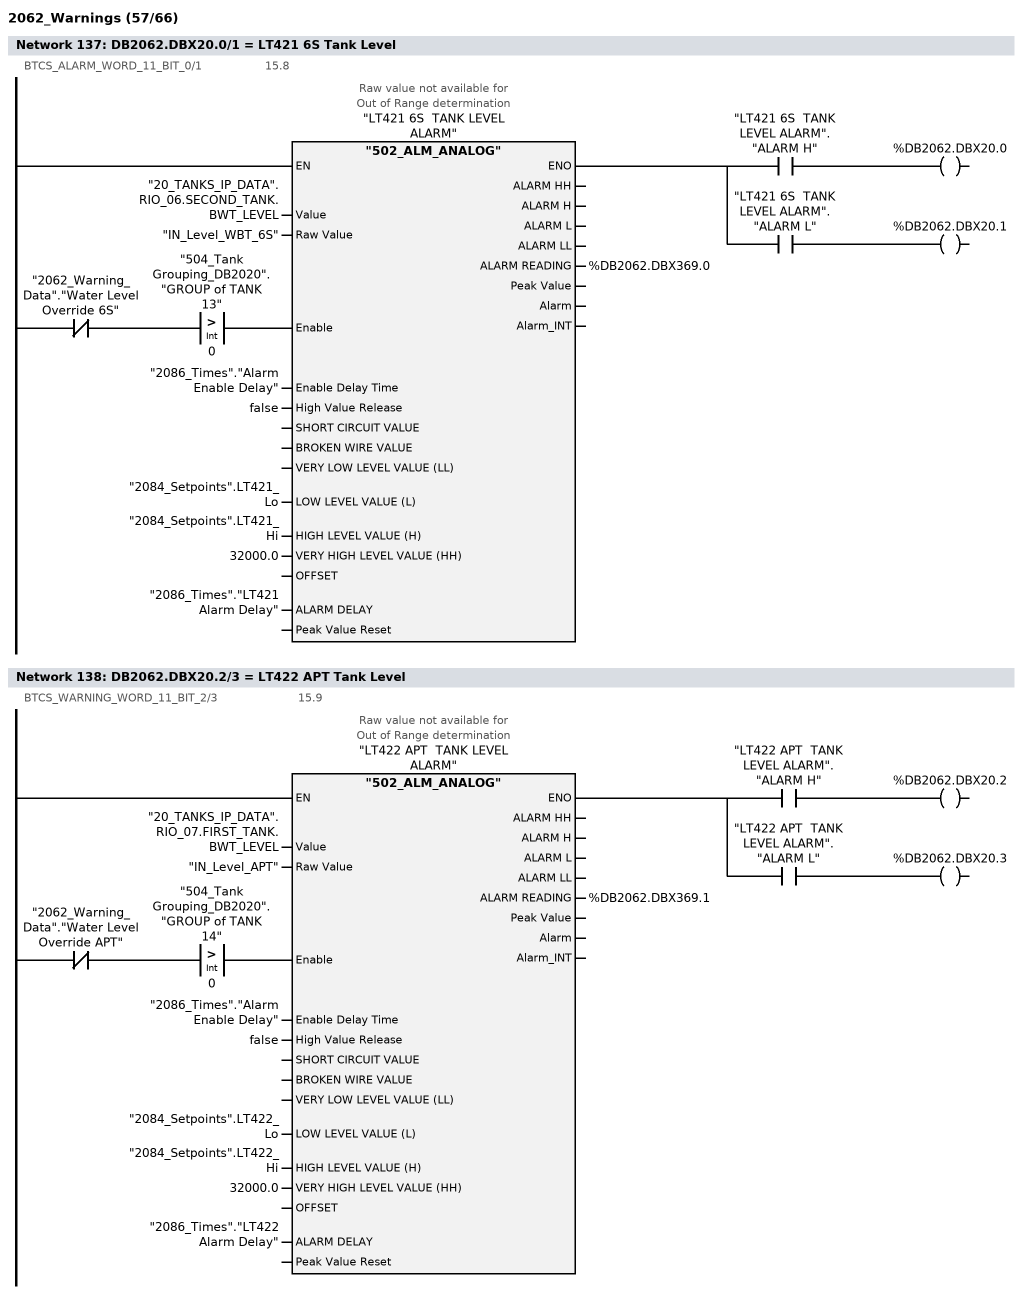
   RUNG wire#powerrail
      "LT421 6S  TANK LEVEL ALARM"(Enable := wire#w1, Value := "20_TANKS_IP_DATA".RIO_06.SECOND_TANK.BWT_LEVEL, "Raw Value" := "IN_Level_WBT_6S", "Enable Delay Time" := "2086_Times"."Alarm Enable Delay", "High Value Release" := false, "SHORT CIRCUIT VALUE" :=, "BROKEN WIRE VALUE" :=, "VERY LOW LEVEL VALUE (LL)" :=, "LOW LEVEL VALUE (L)" := "2084_Setpoints".LT421_Lo, "HIGH LEVEL VALUE (H)" := "2084_Setpoints".LT421_Hi, "VERY HIGH LEVEL VALUE (HH)" := 32000.0, OFFSET :=, "ALARM DELAY" := "2086_Times"."LT421 Alarm Delay", "Peak Value Reset" :=, "ALARM HH" =>, "ALARM H" =>, "ALARM L" =>, "ALARM LL" =>, "ALARM READING" => %DB2062.DBX369.0, "Peak Value" =>, Alarm =>, Alarm_INT =>)   // Raw value not available for Out of Range determination
      wire#w2
      Contact( "LT421 6S  TANK LEVEL ALARM"."ALARM H" )
      Coil( %DB2062.DBX20.0 )
   END_RUNG
   RUNG wire#powerrail
      I_Contact( "2062_Warning_Data"."Water Level Override 6S" )
      { S7_Templates := "SrcType := Int" } GT_Contact(in1 := "504_Tank Grouping_DB2020"."GROUP of TANK 13", in2 := 0)
   END_RUNG wire#w1
   RUNG wire#w2
      Contact( "LT421 6S  TANK LEVEL ALARM"."ALARM L" )
      Coil( %DB2062.DBX20.1 )
   END_RUNG
   // the same network as SCL:
   "LT421 6S  TANK LEVEL ALARM"(Value := "20_TANKS_IP_DATA".RIO_06.SECOND_TANK.BWT_LEVEL,   // "502_ALM_ANALOG": Raw value not available for Out of Range determination
                           "Raw Value" := "IN_Level_WBT_6S",
                           Enable := NOT "2062_Warning_Data"."Water Level Override 6S" AND ("504_Tank Grouping_DB2020"."GROUP of TANK 13" > 0),
                           "Enable Delay Time" := "2086_Times"."Alarm Enable Delay",
                           "High Value Release" := false,
                           "LOW LEVEL VALUE (L)" := "2084_Setpoints".LT421_Lo,
                           "HIGH LEVEL VALUE (H)" := "2084_Setpoints".LT421_Hi,
                           "VERY HIGH LEVEL VALUE (HH)" := 32000.0,
                           "ALARM DELAY" := "2086_Times"."LT421 Alarm Delay",
                           "ALARM READING" => %DB2062.DBX369.0,
                           ENO => #_w1);
   %DB2062.DBX20.0 := #_w1 AND "LT421 6S  TANK LEVEL ALARM"."ALARM H";
   %DB2062.DBX20.1 := #_w1 AND "LT421 6S  TANK LEVEL ALARM"."ALARM L";
END_REGION

REGION Network 138: DB2062.DBX20.2/3 = LT422 APT Tank Level
   // BTCS_WARNING_WORD_11_BIT_2/3                       15.9
   RUNG wire#powerrail
      "LT422 APT  TANK LEVEL ALARM"(Enable := wire#w1, Value := "20_TANKS_IP_DATA".RIO_07.FIRST_TANK.BWT_LEVEL, "Raw Value" := "IN_Level_APT", "Enable Delay Time" := "2086_Times"."Alarm Enable Delay", "High Value Release" := false, "SHORT CIRCUIT VALUE" :=, "BROKEN WIRE VALUE" :=, "VERY LOW LEVEL VALUE (LL)" :=, "LOW LEVEL VALUE (L)" := "2084_Setpoints".LT422_Lo, "HIGH LEVEL VALUE (H)" := "2084_Setpoints".LT422_Hi, "VERY HIGH LEVEL VALUE (HH)" := 32000.0, OFFSET :=, "ALARM DELAY" := "2086_Times"."LT422 Alarm Delay", "Peak Value Reset" :=, "ALARM HH" =>, "ALARM H" =>, "ALARM L" =>, "ALARM LL" =>, "ALARM READING" => %DB2062.DBX369.1, "Peak Value" =>, Alarm =>, Alarm_INT =>)   // Raw value not available for Out of Range determination
      wire#w2
      Contact( "LT422 APT  TANK LEVEL ALARM"."ALARM H" )
      Coil( %DB2062.DBX20.2 )
   END_RUNG
   RUNG wire#powerrail
      I_Contact( "2062_Warning_Data"."Water Level Override APT" )
      { S7_Templates := "SrcType := Int" } GT_Contact(in1 := "504_Tank Grouping_DB2020"."GROUP of TANK 14", in2 := 0)
   END_RUNG wire#w1
   RUNG wire#w2
      Contact( "LT422 APT  TANK LEVEL ALARM"."ALARM L" )
      Coil( %DB2062.DBX20.3 )
   END_RUNG
   // the same network as SCL:
   "LT422 APT  TANK LEVEL ALARM"(Value := "20_TANKS_IP_DATA".RIO_07.FIRST_TANK.BWT_LEVEL,   // "502_ALM_ANALOG": Raw value not available for Out of Range determination
                           "Raw Value" := "IN_Level_APT",
                           Enable := NOT "2062_Warning_Data"."Water Level Override APT" AND ("504_Tank Grouping_DB2020"."GROUP of TANK 14" > 0),
                           "Enable Delay Time" := "2086_Times"."Alarm Enable Delay",
                           "High Value Release" := false,
                           "LOW LEVEL VALUE (L)" := "2084_Setpoints".LT422_Lo,
                           "HIGH LEVEL VALUE (H)" := "2084_Setpoints".LT422_Hi,
                           "VERY HIGH LEVEL VALUE (HH)" := 32000.0,
                           "ALARM DELAY" := "2086_Times"."LT422 Alarm Delay",
                           "ALARM READING" => %DB2062.DBX369.1,
                           ENO => #_w1);
   %DB2062.DBX20.2 := #_w1 AND "LT422 APT  TANK LEVEL ALARM"."ALARM H";
   %DB2062.DBX20.3 := #_w1 AND "LT422 APT  TANK LEVEL ALARM"."ALARM L";
END_REGION

REGION Network 140: Alarm Tank 1
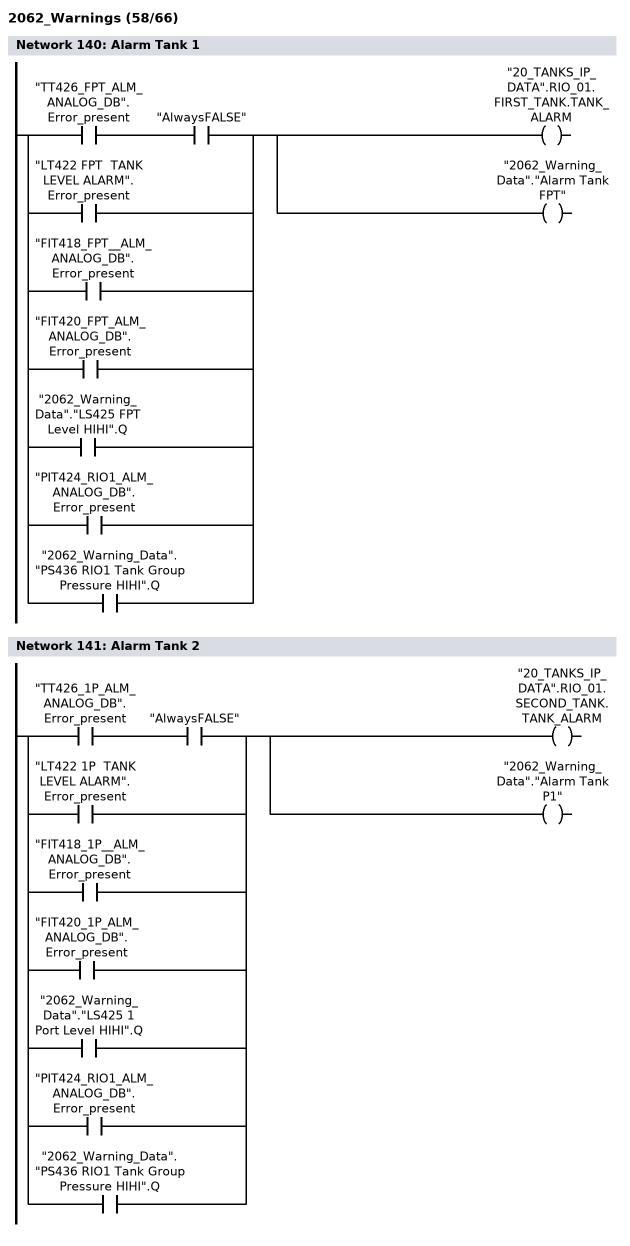
   RUNG wire#powerrail
      Contact( "TT426_FPT_ALM_ANALOG_DB".Error_present )
      Contact( "AlwaysFALSE" )
      wire#w1
      Coil( "20_TANKS_IP_DATA".RIO_01.FIRST_TANK.TANK_ALARM )
   END_RUNG
   RUNG wire#powerrail
      Contact( "LT422 FPT  TANK LEVEL ALARM".Error_present )
   END_RUNG wire#w1
   RUNG wire#powerrail
      Contact( "FIT418_FPT__ALM_ANALOG_DB".Error_present )
   END_RUNG wire#w1
   RUNG wire#powerrail
      Contact( "FIT420_FPT_ALM_ANALOG_DB".Error_present )
   END_RUNG wire#w1
   RUNG wire#powerrail
      Contact( "2062_Warning_Data"."LS425 FPT Level HIHI".Q )
   END_RUNG wire#w1
   RUNG wire#powerrail
      Contact( "PIT424_RIO1_ALM_ANALOG_DB".Error_present )
   END_RUNG wire#w1
   RUNG wire#powerrail
      Contact( "2062_Warning_Data"."PS436 RIO1 Tank Group Pressure HIHI".Q )
   END_RUNG wire#w1
   RUNG wire#w1
      Coil( "2062_Warning_Data"."Alarm Tank FPT" )
   END_RUNG
   // the same network as SCL:
   "20_TANKS_IP_DATA".RIO_01.FIRST_TANK.TANK_ALARM := ("TT426_FPT_ALM_ANALOG_DB".Error_present AND "AlwaysFALSE") OR "LT422 FPT  TANK LEVEL ALARM".Error_present OR "FIT418_FPT__ALM_ANALOG_DB".Error_present OR "FIT420_FPT_ALM_ANALOG_DB".Error_present OR "2062_Warning_Data"."LS425 FPT Level HIHI".Q OR "PIT424_RIO1_ALM_ANALOG_DB".Error_present OR "2062_Warning_Data"."PS436 RIO1 Tank Group Pressure HIHI".Q;
   "2062_Warning_Data"."Alarm Tank FPT" := "20_TANKS_IP_DATA".RIO_01.FIRST_TANK.TANK_ALARM;
END_REGION

REGION Network 141: Alarm Tank 2
   RUNG wire#powerrail
      Contact( "TT426_1P_ALM_ANALOG_DB".Error_present )
      Contact( "AlwaysFALSE" )
      wire#w1
      Coil( "20_TANKS_IP_DATA".RIO_01.SECOND_TANK.TANK_ALARM )
   END_RUNG
   RUNG wire#powerrail
      Contact( "LT422 1P  TANK LEVEL ALARM".Error_present )
   END_RUNG wire#w1
   RUNG wire#powerrail
      Contact( "FIT418_1P__ALM_ANALOG_DB".Error_present )
   END_RUNG wire#w1
   RUNG wire#powerrail
      Contact( "FIT420_1P_ALM_ANALOG_DB".Error_present )
   END_RUNG wire#w1
   RUNG wire#powerrail
      Contact( "2062_Warning_Data"."LS425 1 Port Level HIHI".Q )
   END_RUNG wire#w1
   RUNG wire#powerrail
      Contact( "PIT424_RIO1_ALM_ANALOG_DB".Error_present )
   END_RUNG wire#w1
   RUNG wire#powerrail
      Contact( "2062_Warning_Data"."PS436 RIO1 Tank Group Pressure HIHI".Q )
   END_RUNG wire#w1
   RUNG wire#w1
      Coil( "2062_Warning_Data"."Alarm Tank P1" )
   END_RUNG
   // the same network as SCL:
   "20_TANKS_IP_DATA".RIO_01.SECOND_TANK.TANK_ALARM := ("TT426_1P_ALM_ANALOG_DB".Error_present AND "AlwaysFALSE") OR "LT422 1P  TANK LEVEL ALARM".Error_present OR "FIT418_1P__ALM_ANALOG_DB".Error_present OR "FIT420_1P_ALM_ANALOG_DB".Error_present OR "2062_Warning_Data"."LS425 1 Port Level HIHI".Q OR "PIT424_RIO1_ALM_ANALOG_DB".Error_present OR "2062_Warning_Data"."PS436 RIO1 Tank Group Pressure HIHI".Q;
   "2062_Warning_Data"."Alarm Tank P1" := "20_TANKS_IP_DATA".RIO_01.SECOND_TANK.TANK_ALARM;
END_REGION

REGION Network 142: Alarm Tank 3
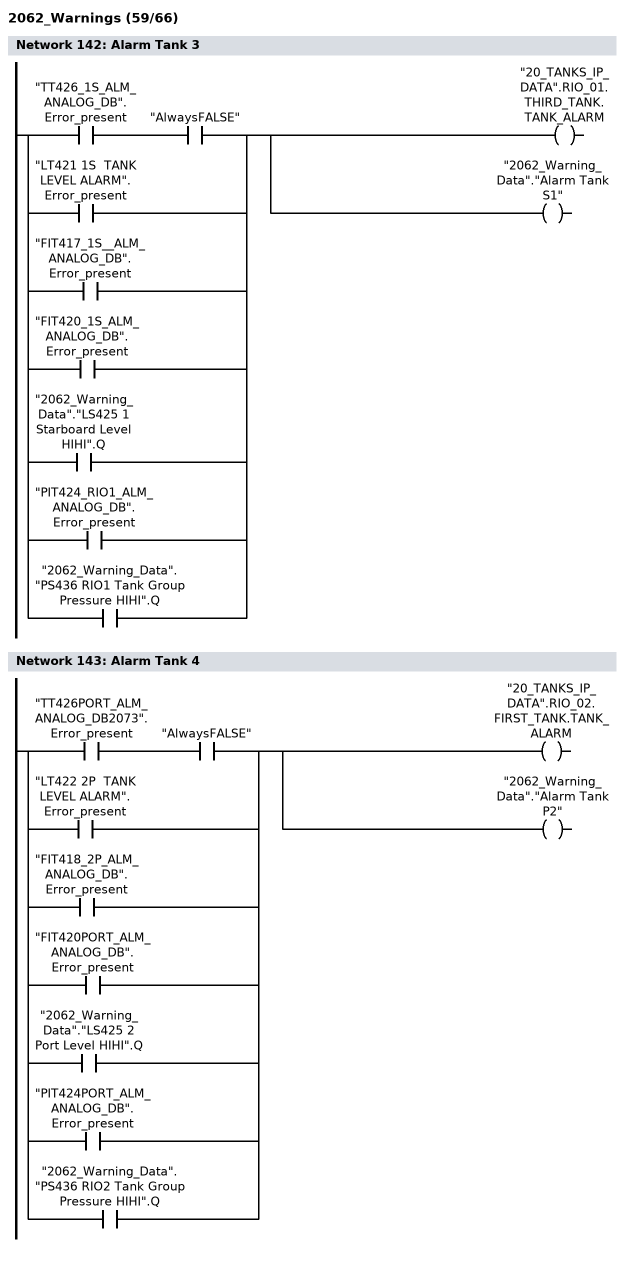
   RUNG wire#powerrail
      Contact( "TT426_1S_ALM_ANALOG_DB".Error_present )
      Contact( "AlwaysFALSE" )
      wire#w1
      Coil( "20_TANKS_IP_DATA".RIO_01.THIRD_TANK.TANK_ALARM )
   END_RUNG
   RUNG wire#powerrail
      Contact( "LT421 1S  TANK LEVEL ALARM".Error_present )
   END_RUNG wire#w1
   RUNG wire#powerrail
      Contact( "FIT417_1S__ALM_ANALOG_DB".Error_present )
   END_RUNG wire#w1
   RUNG wire#powerrail
      Contact( "FIT420_1S_ALM_ANALOG_DB".Error_present )
   END_RUNG wire#w1
   RUNG wire#powerrail
      Contact( "2062_Warning_Data"."LS425 1 Starboard Level HIHI".Q )
   END_RUNG wire#w1
   RUNG wire#powerrail
      Contact( "PIT424_RIO1_ALM_ANALOG_DB".Error_present )
   END_RUNG wire#w1
   RUNG wire#powerrail
      Contact( "2062_Warning_Data"."PS436 RIO1 Tank Group Pressure HIHI".Q )
   END_RUNG wire#w1
   RUNG wire#w1
      Coil( "2062_Warning_Data"."Alarm Tank S1" )
   END_RUNG
   // the same network as SCL:
   "20_TANKS_IP_DATA".RIO_01.THIRD_TANK.TANK_ALARM := ("TT426_1S_ALM_ANALOG_DB".Error_present AND "AlwaysFALSE") OR "LT421 1S  TANK LEVEL ALARM".Error_present OR "FIT417_1S__ALM_ANALOG_DB".Error_present OR "FIT420_1S_ALM_ANALOG_DB".Error_present OR "2062_Warning_Data"."LS425 1 Starboard Level HIHI".Q OR "PIT424_RIO1_ALM_ANALOG_DB".Error_present OR "2062_Warning_Data"."PS436 RIO1 Tank Group Pressure HIHI".Q;
   "2062_Warning_Data"."Alarm Tank S1" := "20_TANKS_IP_DATA".RIO_01.THIRD_TANK.TANK_ALARM;
END_REGION

REGION Network 143: Alarm Tank 4
   RUNG wire#powerrail
      Contact( "TT426PORT_ALM_ANALOG_DB2073".Error_present )
      Contact( "AlwaysFALSE" )
      wire#w1
      Coil( "20_TANKS_IP_DATA".RIO_02.FIRST_TANK.TANK_ALARM )
   END_RUNG
   RUNG wire#powerrail
      Contact( "LT422 2P  TANK LEVEL ALARM".Error_present )
   END_RUNG wire#w1
   RUNG wire#powerrail
      Contact( "FIT418_2P_ALM_ANALOG_DB".Error_present )
   END_RUNG wire#w1
   RUNG wire#powerrail
      Contact( "FIT420PORT_ALM_ANALOG_DB".Error_present )
   END_RUNG wire#w1
   RUNG wire#powerrail
      Contact( "2062_Warning_Data"."LS425 2 Port Level HIHI".Q )
   END_RUNG wire#w1
   RUNG wire#powerrail
      Contact( "PIT424PORT_ALM_ANALOG_DB".Error_present )
   END_RUNG wire#w1
   RUNG wire#powerrail
      Contact( "2062_Warning_Data"."PS436 RIO2 Tank Group Pressure HIHI".Q )
   END_RUNG wire#w1
   RUNG wire#w1
      Coil( "2062_Warning_Data"."Alarm Tank P2" )
   END_RUNG
   // the same network as SCL:
   "20_TANKS_IP_DATA".RIO_02.FIRST_TANK.TANK_ALARM := ("TT426PORT_ALM_ANALOG_DB2073".Error_present AND "AlwaysFALSE") OR "LT422 2P  TANK LEVEL ALARM".Error_present OR "FIT418_2P_ALM_ANALOG_DB".Error_present OR "FIT420PORT_ALM_ANALOG_DB".Error_present OR "2062_Warning_Data"."LS425 2 Port Level HIHI".Q OR "PIT424PORT_ALM_ANALOG_DB".Error_present OR "2062_Warning_Data"."PS436 RIO2 Tank Group Pressure HIHI".Q;
   "2062_Warning_Data"."Alarm Tank P2" := "20_TANKS_IP_DATA".RIO_02.FIRST_TANK.TANK_ALARM;
END_REGION

REGION Network 144: Alarm Tank 5
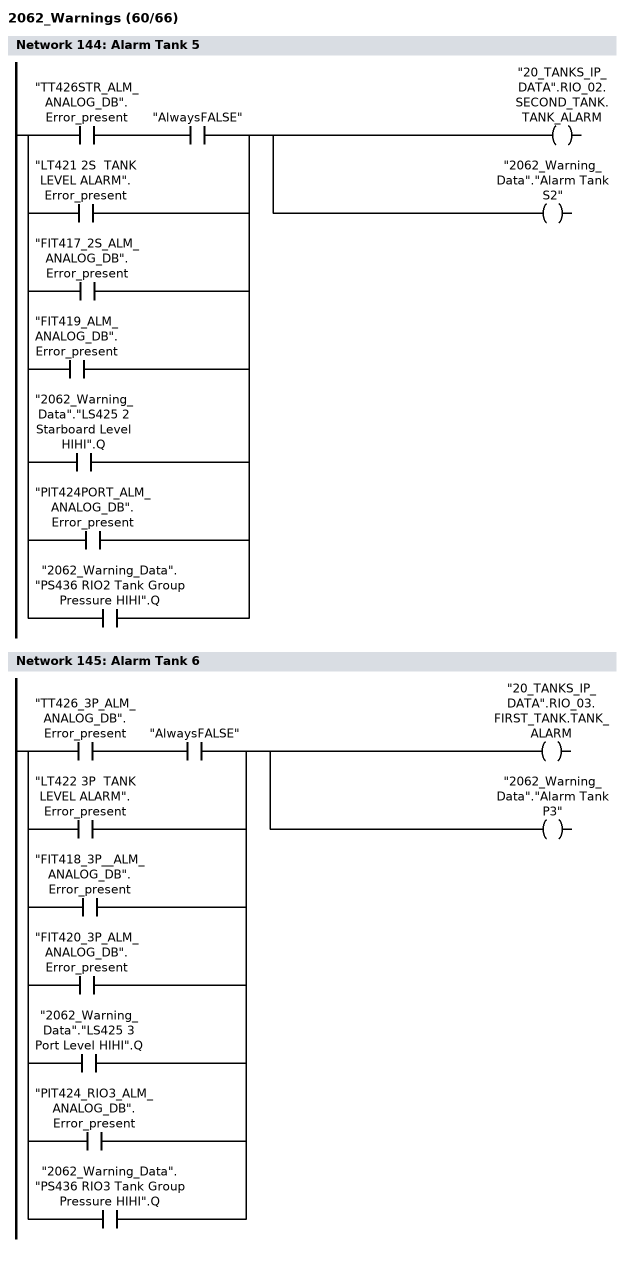
   RUNG wire#powerrail
      Contact( "TT426STR_ALM_ANALOG_DB".Error_present )
      Contact( "AlwaysFALSE" )
      wire#w1
      Coil( "20_TANKS_IP_DATA".RIO_02.SECOND_TANK.TANK_ALARM )
   END_RUNG
   RUNG wire#powerrail
      Contact( "LT421 2S  TANK LEVEL ALARM".Error_present )
   END_RUNG wire#w1
   RUNG wire#powerrail
      Contact( "FIT417_2S_ALM_ANALOG_DB".Error_present )
   END_RUNG wire#w1
   RUNG wire#powerrail
      Contact( "FIT419_ALM_ANALOG_DB".Error_present )
   END_RUNG wire#w1
   RUNG wire#powerrail
      Contact( "2062_Warning_Data"."LS425 2 Starboard Level HIHI".Q )
   END_RUNG wire#w1
   RUNG wire#powerrail
      Contact( "PIT424PORT_ALM_ANALOG_DB".Error_present )
   END_RUNG wire#w1
   RUNG wire#powerrail
      Contact( "2062_Warning_Data"."PS436 RIO2 Tank Group Pressure HIHI".Q )
   END_RUNG wire#w1
   RUNG wire#w1
      Coil( "2062_Warning_Data"."Alarm Tank S2" )
   END_RUNG
   // the same network as SCL:
   "20_TANKS_IP_DATA".RIO_02.SECOND_TANK.TANK_ALARM := ("TT426STR_ALM_ANALOG_DB".Error_present AND "AlwaysFALSE") OR "LT421 2S  TANK LEVEL ALARM".Error_present OR "FIT417_2S_ALM_ANALOG_DB".Error_present OR "FIT419_ALM_ANALOG_DB".Error_present OR "2062_Warning_Data"."LS425 2 Starboard Level HIHI".Q OR "PIT424PORT_ALM_ANALOG_DB".Error_present OR "2062_Warning_Data"."PS436 RIO2 Tank Group Pressure HIHI".Q;
   "2062_Warning_Data"."Alarm Tank S2" := "20_TANKS_IP_DATA".RIO_02.SECOND_TANK.TANK_ALARM;
END_REGION

REGION Network 145: Alarm Tank 6
   RUNG wire#powerrail
      Contact( "TT426_3P_ALM_ANALOG_DB".Error_present )
      Contact( "AlwaysFALSE" )
      wire#w1
      Coil( "20_TANKS_IP_DATA".RIO_03.FIRST_TANK.TANK_ALARM )
   END_RUNG
   RUNG wire#powerrail
      Contact( "LT422 3P  TANK LEVEL ALARM".Error_present )
   END_RUNG wire#w1
   RUNG wire#powerrail
      Contact( "FIT418_3P__ALM_ANALOG_DB".Error_present )
   END_RUNG wire#w1
   RUNG wire#powerrail
      Contact( "FIT420_3P_ALM_ANALOG_DB".Error_present )
   END_RUNG wire#w1
   RUNG wire#powerrail
      Contact( "2062_Warning_Data"."LS425 3 Port Level HIHI".Q )
   END_RUNG wire#w1
   RUNG wire#powerrail
      Contact( "PIT424_RIO3_ALM_ANALOG_DB".Error_present )
   END_RUNG wire#w1
   RUNG wire#powerrail
      Contact( "2062_Warning_Data"."PS436 RIO3 Tank Group Pressure HIHI".Q )
   END_RUNG wire#w1
   RUNG wire#w1
      Coil( "2062_Warning_Data"."Alarm Tank P3" )
   END_RUNG
   // the same network as SCL:
   "20_TANKS_IP_DATA".RIO_03.FIRST_TANK.TANK_ALARM := ("TT426_3P_ALM_ANALOG_DB".Error_present AND "AlwaysFALSE") OR "LT422 3P  TANK LEVEL ALARM".Error_present OR "FIT418_3P__ALM_ANALOG_DB".Error_present OR "FIT420_3P_ALM_ANALOG_DB".Error_present OR "2062_Warning_Data"."LS425 3 Port Level HIHI".Q OR "PIT424_RIO3_ALM_ANALOG_DB".Error_present OR "2062_Warning_Data"."PS436 RIO3 Tank Group Pressure HIHI".Q;
   "2062_Warning_Data"."Alarm Tank P3" := "20_TANKS_IP_DATA".RIO_03.FIRST_TANK.TANK_ALARM;
END_REGION

REGION Network 146: Alarm Tank 7
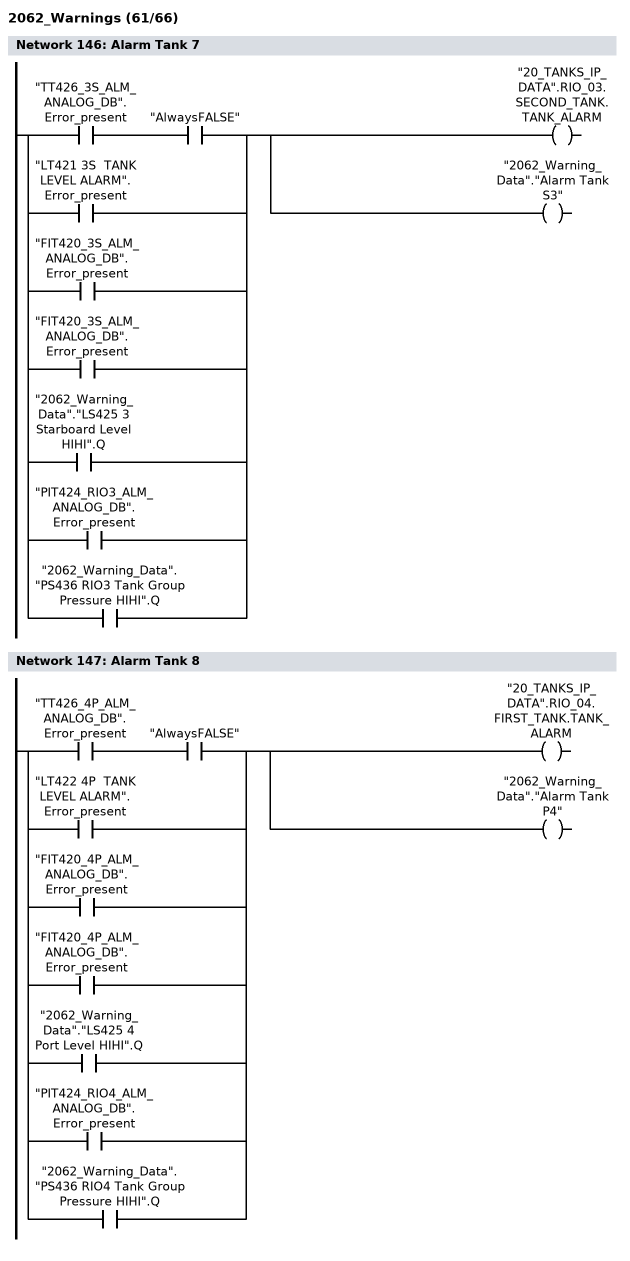
   RUNG wire#powerrail
      Contact( "TT426_3S_ALM_ANALOG_DB".Error_present )
      Contact( "AlwaysFALSE" )
      wire#w1
      Coil( "20_TANKS_IP_DATA".RIO_03.SECOND_TANK.TANK_ALARM )
   END_RUNG
   RUNG wire#powerrail
      Contact( "LT421 3S  TANK LEVEL ALARM".Error_present )
   END_RUNG wire#w1
   RUNG wire#powerrail
      Contact( "FIT420_3S_ALM_ANALOG_DB".Error_present )
   END_RUNG wire#w1
   RUNG wire#powerrail
      Contact( "FIT420_3S_ALM_ANALOG_DB".Error_present )
   END_RUNG wire#w1
   RUNG wire#powerrail
      Contact( "2062_Warning_Data"."LS425 3 Starboard Level HIHI".Q )
   END_RUNG wire#w1
   RUNG wire#powerrail
      Contact( "PIT424_RIO3_ALM_ANALOG_DB".Error_present )
   END_RUNG wire#w1
   RUNG wire#powerrail
      Contact( "2062_Warning_Data"."PS436 RIO3 Tank Group Pressure HIHI".Q )
   END_RUNG wire#w1
   RUNG wire#w1
      Coil( "2062_Warning_Data"."Alarm Tank S3" )
   END_RUNG
   // the same network as SCL:
   "20_TANKS_IP_DATA".RIO_03.SECOND_TANK.TANK_ALARM := ("TT426_3S_ALM_ANALOG_DB".Error_present AND "AlwaysFALSE") OR "LT421 3S  TANK LEVEL ALARM".Error_present OR "FIT420_3S_ALM_ANALOG_DB".Error_present OR "FIT420_3S_ALM_ANALOG_DB".Error_present OR "2062_Warning_Data"."LS425 3 Starboard Level HIHI".Q OR "PIT424_RIO3_ALM_ANALOG_DB".Error_present OR "2062_Warning_Data"."PS436 RIO3 Tank Group Pressure HIHI".Q;
   "2062_Warning_Data"."Alarm Tank S3" := "20_TANKS_IP_DATA".RIO_03.SECOND_TANK.TANK_ALARM;
END_REGION

REGION Network 147: Alarm Tank 8
   RUNG wire#powerrail
      Contact( "TT426_4P_ALM_ANALOG_DB".Error_present )
      Contact( "AlwaysFALSE" )
      wire#w1
      Coil( "20_TANKS_IP_DATA".RIO_04.FIRST_TANK.TANK_ALARM )
   END_RUNG
   RUNG wire#powerrail
      Contact( "LT422 4P  TANK LEVEL ALARM".Error_present )
   END_RUNG wire#w1
   RUNG wire#powerrail
      Contact( "FIT420_4P_ALM_ANALOG_DB".Error_present )
   END_RUNG wire#w1
   RUNG wire#powerrail
      Contact( "FIT420_4P_ALM_ANALOG_DB".Error_present )
   END_RUNG wire#w1
   RUNG wire#powerrail
      Contact( "2062_Warning_Data"."LS425 4 Port Level HIHI".Q )
   END_RUNG wire#w1
   RUNG wire#powerrail
      Contact( "PIT424_RIO4_ALM_ANALOG_DB".Error_present )
   END_RUNG wire#w1
   RUNG wire#powerrail
      Contact( "2062_Warning_Data"."PS436 RIO4 Tank Group Pressure HIHI".Q )
   END_RUNG wire#w1
   RUNG wire#w1
      Coil( "2062_Warning_Data"."Alarm Tank P4" )
   END_RUNG
   // the same network as SCL:
   "20_TANKS_IP_DATA".RIO_04.FIRST_TANK.TANK_ALARM := ("TT426_4P_ALM_ANALOG_DB".Error_present AND "AlwaysFALSE") OR "LT422 4P  TANK LEVEL ALARM".Error_present OR "FIT420_4P_ALM_ANALOG_DB".Error_present OR "FIT420_4P_ALM_ANALOG_DB".Error_present OR "2062_Warning_Data"."LS425 4 Port Level HIHI".Q OR "PIT424_RIO4_ALM_ANALOG_DB".Error_present OR "2062_Warning_Data"."PS436 RIO4 Tank Group Pressure HIHI".Q;
   "2062_Warning_Data"."Alarm Tank P4" := "20_TANKS_IP_DATA".RIO_04.FIRST_TANK.TANK_ALARM;
END_REGION

REGION Network 148: Alarm Tank 9
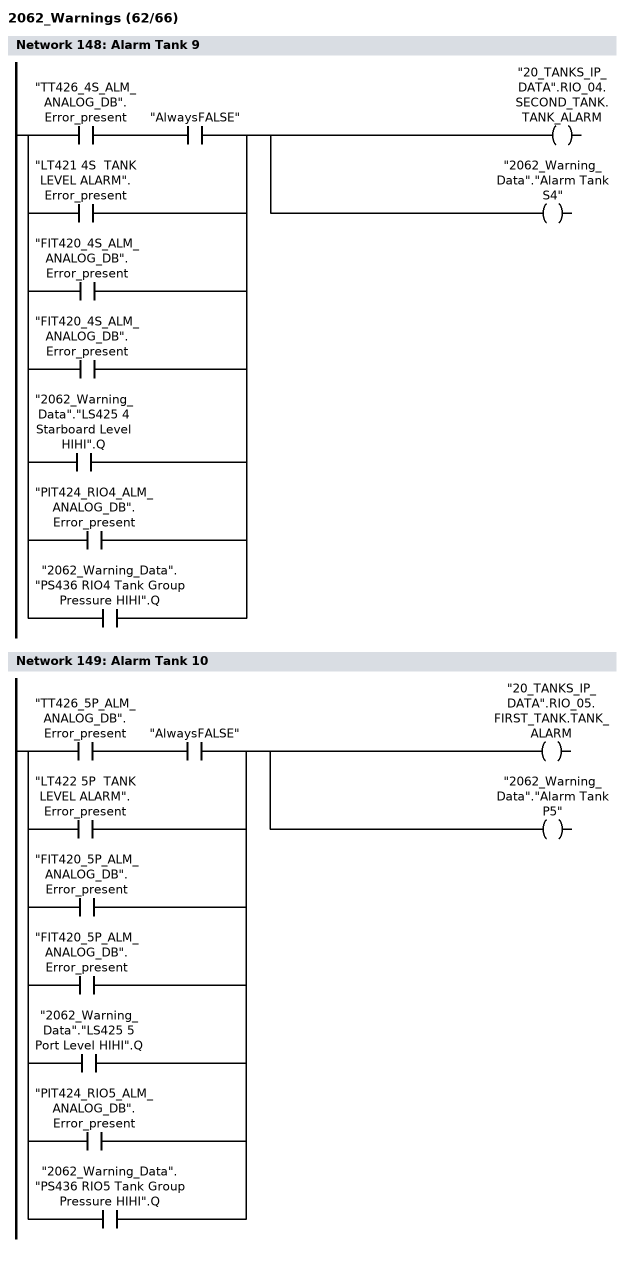
   RUNG wire#powerrail
      Contact( "TT426_4S_ALM_ANALOG_DB".Error_present )
      Contact( "AlwaysFALSE" )
      wire#w1
      Coil( "20_TANKS_IP_DATA".RIO_04.SECOND_TANK.TANK_ALARM )
   END_RUNG
   RUNG wire#powerrail
      Contact( "LT421 4S  TANK LEVEL ALARM".Error_present )
   END_RUNG wire#w1
   RUNG wire#powerrail
      Contact( "FIT420_4S_ALM_ANALOG_DB".Error_present )
   END_RUNG wire#w1
   RUNG wire#powerrail
      Contact( "FIT420_4S_ALM_ANALOG_DB".Error_present )
   END_RUNG wire#w1
   RUNG wire#powerrail
      Contact( "2062_Warning_Data"."LS425 4 Starboard Level HIHI".Q )
   END_RUNG wire#w1
   RUNG wire#powerrail
      Contact( "PIT424_RIO4_ALM_ANALOG_DB".Error_present )
   END_RUNG wire#w1
   RUNG wire#powerrail
      Contact( "2062_Warning_Data"."PS436 RIO4 Tank Group Pressure HIHI".Q )
   END_RUNG wire#w1
   RUNG wire#w1
      Coil( "2062_Warning_Data"."Alarm Tank S4" )
   END_RUNG
   // the same network as SCL:
   "20_TANKS_IP_DATA".RIO_04.SECOND_TANK.TANK_ALARM := ("TT426_4S_ALM_ANALOG_DB".Error_present AND "AlwaysFALSE") OR "LT421 4S  TANK LEVEL ALARM".Error_present OR "FIT420_4S_ALM_ANALOG_DB".Error_present OR "FIT420_4S_ALM_ANALOG_DB".Error_present OR "2062_Warning_Data"."LS425 4 Starboard Level HIHI".Q OR "PIT424_RIO4_ALM_ANALOG_DB".Error_present OR "2062_Warning_Data"."PS436 RIO4 Tank Group Pressure HIHI".Q;
   "2062_Warning_Data"."Alarm Tank S4" := "20_TANKS_IP_DATA".RIO_04.SECOND_TANK.TANK_ALARM;
END_REGION

REGION Network 149: Alarm Tank 10
   RUNG wire#powerrail
      Contact( "TT426_5P_ALM_ANALOG_DB".Error_present )
      Contact( "AlwaysFALSE" )
      wire#w1
      Coil( "20_TANKS_IP_DATA".RIO_05.FIRST_TANK.TANK_ALARM )
   END_RUNG
   RUNG wire#powerrail
      Contact( "LT422 5P  TANK LEVEL ALARM".Error_present )
   END_RUNG wire#w1
   RUNG wire#powerrail
      Contact( "FIT420_5P_ALM_ANALOG_DB".Error_present )
   END_RUNG wire#w1
   RUNG wire#powerrail
      Contact( "FIT420_5P_ALM_ANALOG_DB".Error_present )
   END_RUNG wire#w1
   RUNG wire#powerrail
      Contact( "2062_Warning_Data"."LS425 5 Port Level HIHI".Q )
   END_RUNG wire#w1
   RUNG wire#powerrail
      Contact( "PIT424_RIO5_ALM_ANALOG_DB".Error_present )
   END_RUNG wire#w1
   RUNG wire#powerrail
      Contact( "2062_Warning_Data"."PS436 RIO5 Tank Group Pressure HIHI".Q )
   END_RUNG wire#w1
   RUNG wire#w1
      Coil( "2062_Warning_Data"."Alarm Tank P5" )
   END_RUNG
   // the same network as SCL:
   "20_TANKS_IP_DATA".RIO_05.FIRST_TANK.TANK_ALARM := ("TT426_5P_ALM_ANALOG_DB".Error_present AND "AlwaysFALSE") OR "LT422 5P  TANK LEVEL ALARM".Error_present OR "FIT420_5P_ALM_ANALOG_DB".Error_present OR "FIT420_5P_ALM_ANALOG_DB".Error_present OR "2062_Warning_Data"."LS425 5 Port Level HIHI".Q OR "PIT424_RIO5_ALM_ANALOG_DB".Error_present OR "2062_Warning_Data"."PS436 RIO5 Tank Group Pressure HIHI".Q;
   "2062_Warning_Data"."Alarm Tank P5" := "20_TANKS_IP_DATA".RIO_05.FIRST_TANK.TANK_ALARM;
END_REGION

REGION Network 150: Alarm Tank 11
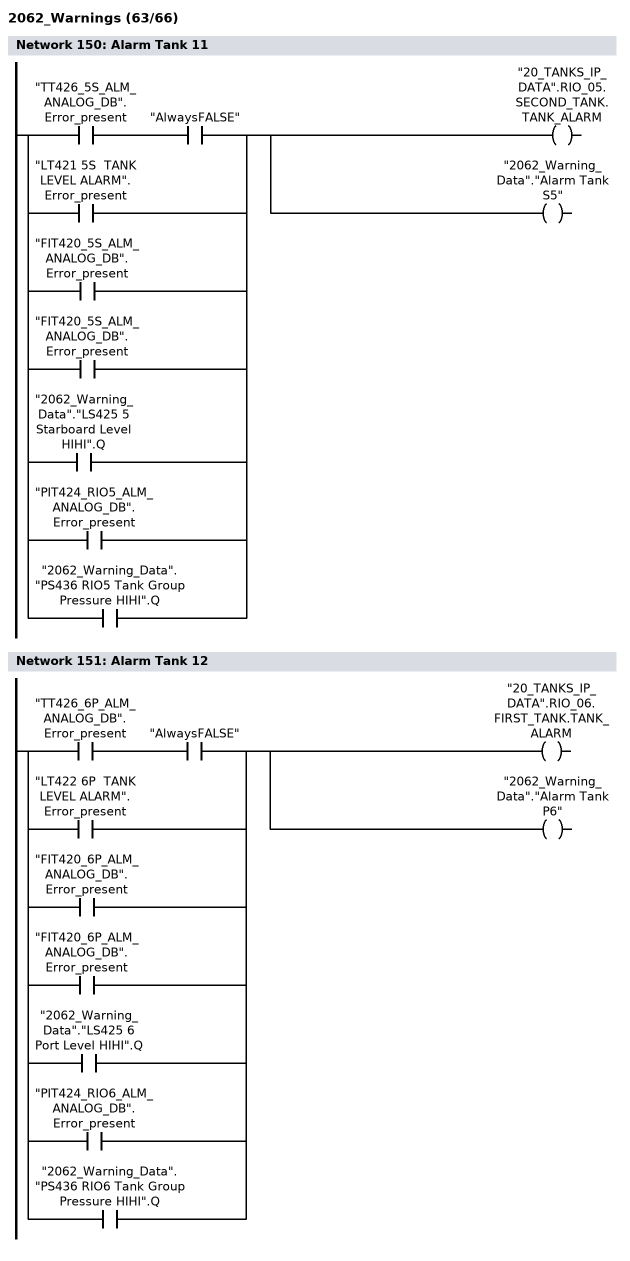
   RUNG wire#powerrail
      Contact( "TT426_5S_ALM_ANALOG_DB".Error_present )
      Contact( "AlwaysFALSE" )
      wire#w1
      Coil( "20_TANKS_IP_DATA".RIO_05.SECOND_TANK.TANK_ALARM )
   END_RUNG
   RUNG wire#powerrail
      Contact( "LT421 5S  TANK LEVEL ALARM".Error_present )
   END_RUNG wire#w1
   RUNG wire#powerrail
      Contact( "FIT420_5S_ALM_ANALOG_DB".Error_present )
   END_RUNG wire#w1
   RUNG wire#powerrail
      Contact( "FIT420_5S_ALM_ANALOG_DB".Error_present )
   END_RUNG wire#w1
   RUNG wire#powerrail
      Contact( "2062_Warning_Data"."LS425 5 Starboard Level HIHI".Q )
   END_RUNG wire#w1
   RUNG wire#powerrail
      Contact( "PIT424_RIO5_ALM_ANALOG_DB".Error_present )
   END_RUNG wire#w1
   RUNG wire#powerrail
      Contact( "2062_Warning_Data"."PS436 RIO5 Tank Group Pressure HIHI".Q )
   END_RUNG wire#w1
   RUNG wire#w1
      Coil( "2062_Warning_Data"."Alarm Tank S5" )
   END_RUNG
   // the same network as SCL:
   "20_TANKS_IP_DATA".RIO_05.SECOND_TANK.TANK_ALARM := ("TT426_5S_ALM_ANALOG_DB".Error_present AND "AlwaysFALSE") OR "LT421 5S  TANK LEVEL ALARM".Error_present OR "FIT420_5S_ALM_ANALOG_DB".Error_present OR "FIT420_5S_ALM_ANALOG_DB".Error_present OR "2062_Warning_Data"."LS425 5 Starboard Level HIHI".Q OR "PIT424_RIO5_ALM_ANALOG_DB".Error_present OR "2062_Warning_Data"."PS436 RIO5 Tank Group Pressure HIHI".Q;
   "2062_Warning_Data"."Alarm Tank S5" := "20_TANKS_IP_DATA".RIO_05.SECOND_TANK.TANK_ALARM;
END_REGION

REGION Network 151: Alarm Tank 12
   RUNG wire#powerrail
      Contact( "TT426_6P_ALM_ANALOG_DB".Error_present )
      Contact( "AlwaysFALSE" )
      wire#w1
      Coil( "20_TANKS_IP_DATA".RIO_06.FIRST_TANK.TANK_ALARM )
   END_RUNG
   RUNG wire#powerrail
      Contact( "LT422 6P  TANK LEVEL ALARM".Error_present )
   END_RUNG wire#w1
   RUNG wire#powerrail
      Contact( "FIT420_6P_ALM_ANALOG_DB".Error_present )
   END_RUNG wire#w1
   RUNG wire#powerrail
      Contact( "FIT420_6P_ALM_ANALOG_DB".Error_present )
   END_RUNG wire#w1
   RUNG wire#powerrail
      Contact( "2062_Warning_Data"."LS425 6 Port Level HIHI".Q )
   END_RUNG wire#w1
   RUNG wire#powerrail
      Contact( "PIT424_RIO6_ALM_ANALOG_DB".Error_present )
   END_RUNG wire#w1
   RUNG wire#powerrail
      Contact( "2062_Warning_Data"."PS436 RIO6 Tank Group Pressure HIHI".Q )
   END_RUNG wire#w1
   RUNG wire#w1
      Coil( "2062_Warning_Data"."Alarm Tank P6" )
   END_RUNG
   // the same network as SCL:
   "20_TANKS_IP_DATA".RIO_06.FIRST_TANK.TANK_ALARM := ("TT426_6P_ALM_ANALOG_DB".Error_present AND "AlwaysFALSE") OR "LT422 6P  TANK LEVEL ALARM".Error_present OR "FIT420_6P_ALM_ANALOG_DB".Error_present OR "FIT420_6P_ALM_ANALOG_DB".Error_present OR "2062_Warning_Data"."LS425 6 Port Level HIHI".Q OR "PIT424_RIO6_ALM_ANALOG_DB".Error_present OR "2062_Warning_Data"."PS436 RIO6 Tank Group Pressure HIHI".Q;
   "2062_Warning_Data"."Alarm Tank P6" := "20_TANKS_IP_DATA".RIO_06.FIRST_TANK.TANK_ALARM;
END_REGION

REGION Network 152: Alarm Tank 13
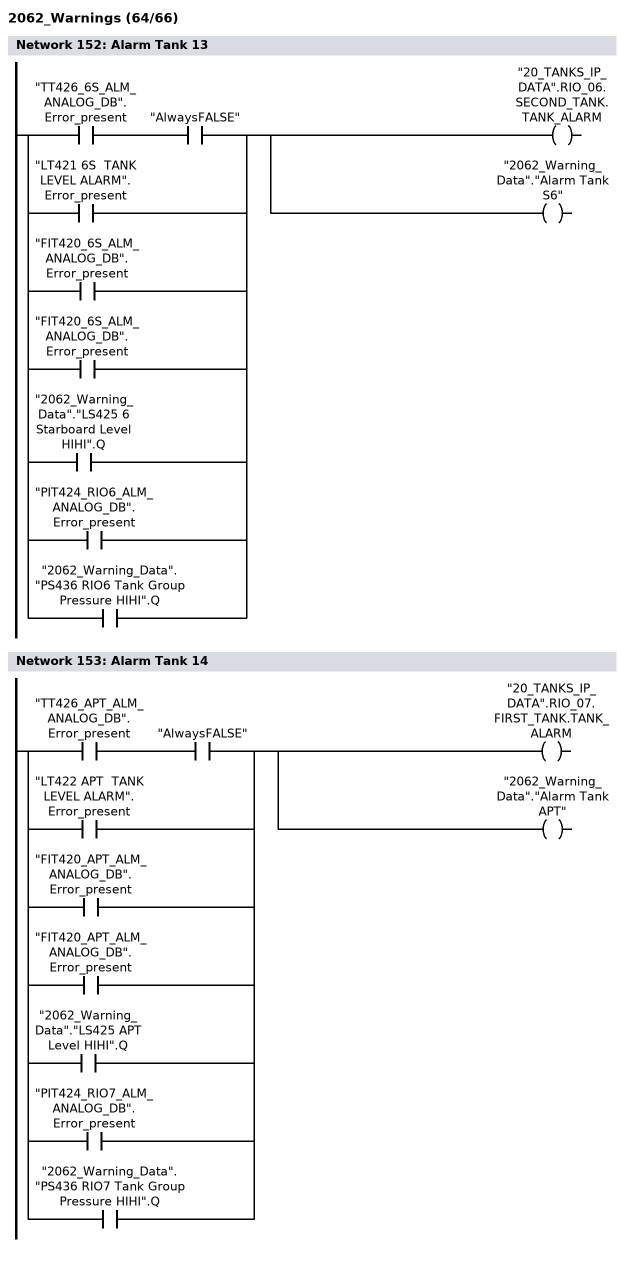
   RUNG wire#powerrail
      Contact( "TT426_6S_ALM_ANALOG_DB".Error_present )
      Contact( "AlwaysFALSE" )
      wire#w1
      Coil( "20_TANKS_IP_DATA".RIO_06.SECOND_TANK.TANK_ALARM )
   END_RUNG
   RUNG wire#powerrail
      Contact( "LT421 6S  TANK LEVEL ALARM".Error_present )
   END_RUNG wire#w1
   RUNG wire#powerrail
      Contact( "FIT420_6S_ALM_ANALOG_DB".Error_present )
   END_RUNG wire#w1
   RUNG wire#powerrail
      Contact( "FIT420_6S_ALM_ANALOG_DB".Error_present )
   END_RUNG wire#w1
   RUNG wire#powerrail
      Contact( "2062_Warning_Data"."LS425 6 Starboard Level HIHI".Q )
   END_RUNG wire#w1
   RUNG wire#powerrail
      Contact( "PIT424_RIO6_ALM_ANALOG_DB".Error_present )
   END_RUNG wire#w1
   RUNG wire#powerrail
      Contact( "2062_Warning_Data"."PS436 RIO6 Tank Group Pressure HIHI".Q )
   END_RUNG wire#w1
   RUNG wire#w1
      Coil( "2062_Warning_Data"."Alarm Tank S6" )
   END_RUNG
   // the same network as SCL:
   "20_TANKS_IP_DATA".RIO_06.SECOND_TANK.TANK_ALARM := ("TT426_6S_ALM_ANALOG_DB".Error_present AND "AlwaysFALSE") OR "LT421 6S  TANK LEVEL ALARM".Error_present OR "FIT420_6S_ALM_ANALOG_DB".Error_present OR "FIT420_6S_ALM_ANALOG_DB".Error_present OR "2062_Warning_Data"."LS425 6 Starboard Level HIHI".Q OR "PIT424_RIO6_ALM_ANALOG_DB".Error_present OR "2062_Warning_Data"."PS436 RIO6 Tank Group Pressure HIHI".Q;
   "2062_Warning_Data"."Alarm Tank S6" := "20_TANKS_IP_DATA".RIO_06.SECOND_TANK.TANK_ALARM;
END_REGION

REGION Network 153: Alarm Tank 14
   RUNG wire#powerrail
      Contact( "TT426_APT_ALM_ANALOG_DB".Error_present )
      Contact( "AlwaysFALSE" )
      wire#w1
      Coil( "20_TANKS_IP_DATA".RIO_07.FIRST_TANK.TANK_ALARM )
   END_RUNG
   RUNG wire#powerrail
      Contact( "LT422 APT  TANK LEVEL ALARM".Error_present )
   END_RUNG wire#w1
   RUNG wire#powerrail
      Contact( "FIT420_APT_ALM_ANALOG_DB".Error_present )
   END_RUNG wire#w1
   RUNG wire#powerrail
      Contact( "FIT420_APT_ALM_ANALOG_DB".Error_present )
   END_RUNG wire#w1
   RUNG wire#powerrail
      Contact( "2062_Warning_Data"."LS425 APT Level HIHI".Q )
   END_RUNG wire#w1
   RUNG wire#powerrail
      Contact( "PIT424_RIO7_ALM_ANALOG_DB".Error_present )
   END_RUNG wire#w1
   RUNG wire#powerrail
      Contact( "2062_Warning_Data"."PS436 RIO7 Tank Group Pressure HIHI".Q )
   END_RUNG wire#w1
   RUNG wire#w1
      Coil( "2062_Warning_Data"."Alarm Tank APT" )
   END_RUNG
   // the same network as SCL:
   "20_TANKS_IP_DATA".RIO_07.FIRST_TANK.TANK_ALARM := ("TT426_APT_ALM_ANALOG_DB".Error_present AND "AlwaysFALSE") OR "LT422 APT  TANK LEVEL ALARM".Error_present OR "FIT420_APT_ALM_ANALOG_DB".Error_present OR "FIT420_APT_ALM_ANALOG_DB".Error_present OR "2062_Warning_Data"."LS425 APT Level HIHI".Q OR "PIT424_RIO7_ALM_ANALOG_DB".Error_present OR "2062_Warning_Data"."PS436 RIO7 Tank Group Pressure HIHI".Q;
   "2062_Warning_Data"."Alarm Tank APT" := "20_TANKS_IP_DATA".RIO_07.FIRST_TANK.TANK_ALARM;
END_REGION

REGION Network 155: New Warning
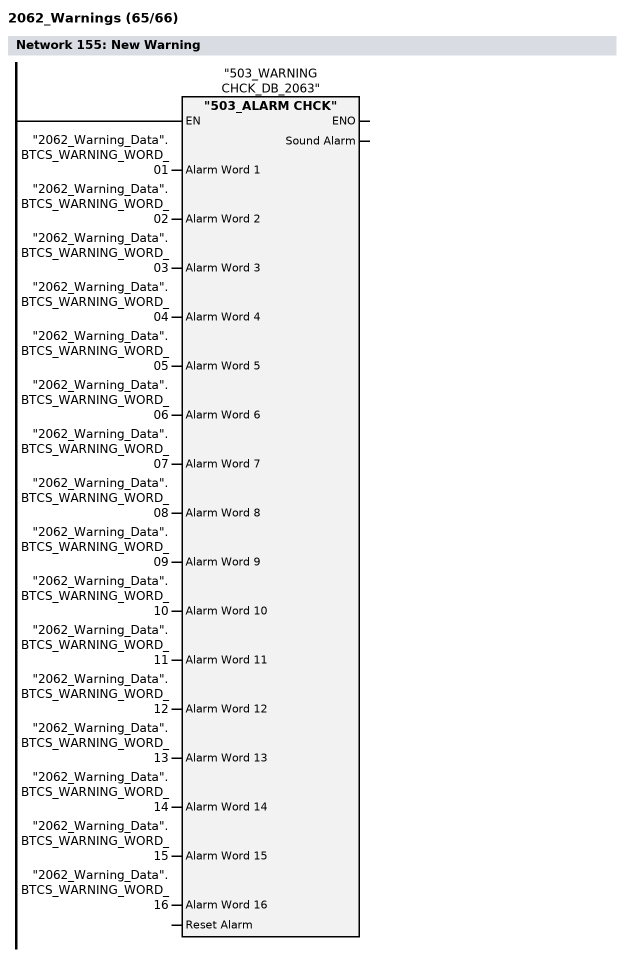
   RUNG wire#powerrail
      "503_WARNING CHCK_DB_2063"("Alarm Word 1" := "2062_Warning_Data".BTCS_WARNING_WORD_01, "Alarm Word 2" := "2062_Warning_Data".BTCS_WARNING_WORD_02, "Alarm Word 3" := "2062_Warning_Data".BTCS_WARNING_WORD_03, "Alarm Word 4" := "2062_Warning_Data".BTCS_WARNING_WORD_04, "Alarm Word 5" := "2062_Warning_Data".BTCS_WARNING_WORD_05, "Alarm Word 6" := "2062_Warning_Data".BTCS_WARNING_WORD_06, "Alarm Word 7" := "2062_Warning_Data".BTCS_WARNING_WORD_07, "Alarm Word 8" := "2062_Warning_Data".BTCS_WARNING_WORD_08, "Alarm Word 9" := "2062_Warning_Data".BTCS_WARNING_WORD_09, "Alarm Word 10" := "2062_Warning_Data".BTCS_WARNING_WORD_10, "Alarm Word 11" := "2062_Warning_Data".BTCS_WARNING_WORD_11, "Alarm Word 12" := "2062_Warning_Data".BTCS_WARNING_WORD_12, "Alarm Word 13" := "2062_Warning_Data".BTCS_WARNING_WORD_13, "Alarm Word 14" := "2062_Warning_Data".BTCS_WARNING_WORD_14, "Alarm Word 15" := "2062_Warning_Data".BTCS_WARNING_WORD_15, "Alarm Word 16" := "2062_Warning_Data".BTCS_WARNING_WORD_16, "Reset Alarm" :=, "Sound Alarm" =>)
   END_RUNG
   // the same network as SCL:
   "503_WARNING CHCK_DB_2063"("Alarm Word 1" := "2062_Warning_Data".BTCS_WARNING_WORD_01,   // "503_ALARM CHCK"
                           "Alarm Word 2" := "2062_Warning_Data".BTCS_WARNING_WORD_02,
                           "Alarm Word 3" := "2062_Warning_Data".BTCS_WARNING_WORD_03,
                           "Alarm Word 4" := "2062_Warning_Data".BTCS_WARNING_WORD_04,
                           "Alarm Word 5" := "2062_Warning_Data".BTCS_WARNING_WORD_05,
                           "Alarm Word 6" := "2062_Warning_Data".BTCS_WARNING_WORD_06,
                           "Alarm Word 7" := "2062_Warning_Data".BTCS_WARNING_WORD_07,
                           "Alarm Word 8" := "2062_Warning_Data".BTCS_WARNING_WORD_08,
                           "Alarm Word 9" := "2062_Warning_Data".BTCS_WARNING_WORD_09,
                           "Alarm Word 10" := "2062_Warning_Data".BTCS_WARNING_WORD_10,
                           "Alarm Word 11" := "2062_Warning_Data".BTCS_WARNING_WORD_11,
                           "Alarm Word 12" := "2062_Warning_Data".BTCS_WARNING_WORD_12,
                           "Alarm Word 13" := "2062_Warning_Data".BTCS_WARNING_WORD_13,
                           "Alarm Word 14" := "2062_Warning_Data".BTCS_WARNING_WORD_14,
                           "Alarm Word 15" := "2062_Warning_Data".BTCS_WARNING_WORD_15,
                           "Alarm Word 16" := "2062_Warning_Data".BTCS_WARNING_WORD_16);
END_REGION

REGION Network 156: Warning Present
